// TIA Portal project "1215C_BREAKOUT_BOARD_IO-LINK_TEMPERATURE" (V19)

(* hardware
DEVICE "BREAKOUT_BOARD_PLC"  S7-1200 Station
   slot 0: "Rack_0"  S7-1200 Rack  Rack  V1.0
   slot 1: "BREAKOUT_BOARD_PLC"  CPU 1215C DC/DC/DC  6ES7 215-1AG40-0XB0  V4.6
DEVICE "BREAKOUT_BOARD_HMI"  KTP400 Basic PN
   slot 0: "BREAKOUT_BOARD_HMI"  KTP400 Basic PN  6AV2 123-2DB03-0AX0  16.0.0.0
   slot 1: "HMI_RT_1"  KTP400 Basic PN  6AV2 123-2DB03-0AX0  16.0.0.0
   slot 5: "BREAKOUT_BOARD_HMI.IE_CP_1"  PROFINET Interface  16.0.0.0
      slot 1: "PROFINET Interface"  PROFINET Interface
         slot 1: "Port_1"  Port
DEVICE "IFM_IO-LINK_MASTER"  GSD.Device.PN
   slot 0: "Rack"  Rack  V1.0
   slot 0: "AL1100"  AL1100  AL1100
      slot 0: "AL1100"  AL1100
      slot 1: "X1"  X1
         slot 1: "Port 1"  Port 1
         slot 2: "Port 2"  Port 2
      slot 1: "4 Ports_1"  4 Ports  AL1100
         slot 0: "IO-Link Master"  IO-Link Master
   slot 1: "IFM ITA2105 IO-Link In  2 Byte + PQI"  IO-Link In  2 Byte + PQI
   slot 2: "Disabled_P2"  Disabled
   slot 3: "Disabled_P3"  Disabled
   slot 4: "Disabled_P4"  Disabled
DEVICE "SCALANCE XB008"  SCALANCE X-Station
   slot 0: "SCALANCE X rack"  Rail
   slot 0: "8PORT_SWITCH"  6GK5 008-0BA10-1AB2  V1.0
*)

// ===== PLC "BREAKOUT_BOARD_PLC"  CPU 1215C DC/DC/DC =====

VAR_GLOBAL   // PLC tag table "PLC_Outputs"
   "DQ0.0" AT %Q0.0 : Bool;   // Digital Output
   "DQ0.1" AT %Q0.1 : Bool;   // Digital Output
   "DQ0.2" AT %Q0.2 : Bool;   // Digital Output
   "DQ0.3" AT %Q0.3 : Bool;   // Digital Output
   "DQ0.4" AT %Q0.4 : Bool;   // Digital Output
   "DQ0.5" AT %Q0.5 : Bool;   // Digital Output
   "DQ0.6" AT %Q0.6 : Bool;   // Digital Output
   "DQ0.7" AT %Q0.7 : Bool;   // Digital Output
   "DQ1.0" AT %Q1.0 : Bool;   // Digital Output
   "DQ1.1" AT %Q1.1 : Bool;   // Digital Output
   "AQ0.0" AT %QW64 : Word;   // Analog Output
   "AQ0.1" AT %QW66 : Word;   // Analog Output
END_VAR

VAR_GLOBAL   // PLC tag table "PLC_Inputs"
   "DI0.0" AT %I0.0 : Bool;   // Digital Input
   "DI0.1" AT %I0.1 : Bool;   // Digital Input
   "DI0.2" AT %I0.2 : Bool;   // Digital Input
   "DI0.3" AT %I0.3 : Bool;   // Digital Input
   "DI0.4" AT %I0.4 : Bool;   // Digital Input
   "DI0.5" AT %I0.5 : Bool;   // Digital Input
   "DI0.6" AT %I0.6 : Bool;   // Digital Input
   "DI0.7" AT %I0.7 : Bool;   // Digital Input
   "DI1.0" AT %I1.0 : Bool;   // Digital Input
   "DI1.1" AT %I1.1 : Bool;   // Digital Input
   "DI1.2" AT %I1.2 : Bool;   // Digital Input
   "DI1.3" AT %I1.3 : Bool;   // Digital Input
   "DI1.4" AT %I1.4 : Bool;   // Digital Input
   "DI1.5" AT %I1.5 : Bool;   // Digital Input
   "AI0.0" AT %IW64 : Word;   // Analog Input
   "AI0.1" AT %IW66 : Word;   // Analog Input
END_VAR

VAR_GLOBAL   // PLC tag table "System_Tags"
   "Clock_Byte" AT %MB0 : Byte;
   "Clock_10Hz" AT %M0.0 : Bool;
   "Clock_5Hz" AT %M0.1 : Bool;
   "Clock_2.5Hz" AT %M0.2 : Bool;
   "Clock_2Hz" AT %M0.3 : Bool;
   "Clock_1.25Hz" AT %M0.4 : Bool;
   "Clock_1Hz" AT %M0.5 : Bool;
   "Clock_0.625Hz" AT %M0.6 : Bool;
   "Clock_0.5Hz" AT %M0.7 : Bool;
   "System_Byte" AT %MB1 : Byte;
   "FirstScan" AT %M1.0 : Bool;
   "DiagStatusUpdate" AT %M1.1 : Bool;
   "AlwaysTRUE" AT %M1.2 : Bool;
   "AlwaysFALSE" AT %M1.3 : Bool;
END_VAR

VAR_GLOBAL   // PLC tag table "Trigger_Tags"
   "xAQ_Trig" AT %M2.0 : Bool;
   "xTrig2" AT %M2.1 : Bool;
   "xTrig3" AT %M2.2 : Bool;
   "xTrig4" AT %M2.3 : Bool;
   "xTrig5" AT %M2.4 : Bool;
END_VAR

VAR_GLOBAL   // PLC tag table "IO-Link_Tags"
   "IFM_TA2105_Temp" AT %IW68 : Int;   // IO-Link Master X1
END_VAR

// folder: WS01_TVET_Workstation/00-I/O_Mapping

DATA_BLOCK "DB001-PLC_I/O"   // DB1
TITLE = PLC I/O Global Database
{ S7_Optimized_Access := 'TRUE' }
VERSION : 0.1
// Variables used to mirror the physical PLC I/O states.
   VAR
      Inputs : Struct   // PLC Inputs Structure
         "xDI0.0" : Bool;
         "xDI0.1" : Bool;
         "xDI0.2" : Bool;
         "xDI0.3" : Bool;
         "xDI0.4" : Bool;
         "xDI0.5" : Bool;
         "xDI0.6" : Bool;
         "xDI0.7" : Bool;
         "xDI1.0" : Bool;
         "xDI1.1" : Bool;
         "xDI1.2" : Bool;
         "xDI1.3" : Bool;
         "xDI1.4" : Bool;
         "xDI1.5" : Bool;
         "rAI0.0_Scaled" : Real;   // 0 to 24648 = 0 to 10 V
         "rAI0.1_Scaled" : Real;   // 0 to 24648 = 0 to 10 V
      END_STRUCT;
      Outputs : Struct   // PLC Outputs Structure
         "xDQ0.0" : Bool;
         "xDQ0.1" : Bool;
         "xDQ0.2" : Bool;
         "xDQ0.3" : Bool;
         "xDQ0.4" : Bool;
         "xDQ0.5" : Bool;
         "xDQ0.6" : Bool;
         "xDQ0.7" : Bool;
         "xDQ1.0" : Bool;
         "xDQ1.1" : Bool;
         "iAQ0.0_RAW" : Int := 0;
         "rAQ0.0_Scaled" : Real;   // 0 to 24648 = 0 to 20 mA
         "iAQ0.1_RAW" : Int := 0;
         "rAQ0.1_Scaled" : Real;   // 0 to 24648 = 0 to 20 mA
      END_STRUCT;
   END_VAR
BEGIN
END_DATA_BLOCK

DATA_BLOCK "DB003-IO-Link_I/O"   // DB3
TITLE = IO-Link I/O Global Database
{ S7_Optimized_Access := 'TRUE' }
VERSION : 0.1
// Variables used to mirror the physical IO-Link I/O states.
   VAR
      Inputs : Struct   // IO-Link Inputs Structure
         wTemp_RAW : Word;   // Temperature Sensor Scaled Value
      END_STRUCT;
      Outputs : Struct   // IO-Link Outputs Structure
         wReserved : Word;
      END_STRUCT;
   END_VAR
BEGIN
END_DATA_BLOCK

// folder: WS01_TVET_Workstation/01-Date_Time

DATA_BLOCK "DB002-DateTime"   // DB2
TITLE = PLC Date/Time Global Database
{ S7_Optimized_Access := 'TRUE' }
VERSION : 0.1
// Variables used to store the PLC date/time & custom date/time formatting.
   VAR
      RD_LOC_T_Ret : Int := 0;   // Return value for Read Local Time Block
      LOCAL_DTL : DTL := DTL#1970-01-01-00:00:00;   // RAW DTL
      "Date" : Date := D#1990-01-01;   // RAW Date
      "Time" : Time_Of_Day := TOD#00:00:00;   // RAW Time
      DTLtoString_Ret : String;   // Return value for DTL to String Block
      sCustomDate_YY : String := '';   // Custom year
      sCustomDate_MM : String := '';   // Custom month
      sCustomDate_DD : String := '';   // Custom Day
      sCustomTime_HH : String := '';   // Custom hour
      sCustomTime_MM : String := '';   // Custom minute
      sCustomDate_DDMMYY : String := '';   // Custom date format
      sCustomTime_HHMM : String := '';   // Custom time format
   END_VAR
BEGIN
END_DATA_BLOCK

// folder: WS01_TVET_Workstation/02-IOLink_Control

DATA_BLOCK "DB004-IOLink_Data"   // DB4
TITLE = IO-Link Data Global Database
{ S7_Optimized_Access := 'TRUE' }
VERSION : 0.1
// Variables used to process data from connected devices.
   VAR
      TempSensor_Data : Struct   // Temperature Sensor Data Structure
         rDeg_C : Real;   // Degrees Celsius
         rDeg_F : Real;   // Degrees Fahrenheit
      END_STRUCT;
   END_VAR
BEGIN
END_DATA_BLOCK

// folder: (top level)

ORGANIZATION_BLOCK "Main"   // OB1, LAD, ProgramCycle
TITLE = "Main Program Sweep (Cycle)"
{ S7_Optimized_Access := 'TRUE' }
VERSION : 0.1
   VAR_INPUT
      Initial_Call : Bool;   // Initial call of this OB
      Remanence : Bool;   // =True, if remanent data are available
   END_VAR
BEGIN

REGION Network 1 (SCL): ================= PROGRAM_INFORMATION =================
   (*
   ==================================================================
   ********************* PLC I/O BREAKOUT BOARD *********************
   ==================================================================

   TVET Workstation WS01:
   1215C DC/DC/DC - 6ES7215-1AG40-0XB0 - IP: 192.168.0.175/24

   KTP400 HMI - 6AV2123-2DB03-0AX0 - IP: 192.168.0.176/24

   IFM IO-Link Master - AL1100 - IP: 192.168.0.177/24

   =======================================================================

   The program has 3 main sections:
   - Date/Time Handler,
   - I/O Handlers,
   - IO-Link Devices Handler.

   Date/Time Handler FC:
   - local PLC date/time is read & formatted into a 24HR time & DD/MM/YYYY.

   I/O Handler FCs:
   - maps the physical PLC inputs & outputs to corresponding tags in DB001,
   - handles scaling of the PLC Analog I/O,
   - maps the IO-Link inputs & outputs to corresponding tags in DB003,
   - ensures that physical I/O tags are only used once in the code.

   IO-Link Device Handler FCs:
   - connected IO-Link devices are controlled in this section with the
     temperature sensor conversion logic being handled by an IFM provided
     FC which scales the input value & converts to Fahrenheit.
   - create & call new FC's for any additional IO-Link devices that may
     get added.

   Additional Notes:
   PLC Tags grouped according to their use/function.

   =======================================================================

   Analog Input Technical data:
   - Number of inputs: 2
   - Type: Voltage (single-ended)
   - Full-scale range: 0 to 10 V
   - Full-scale range (data word): 0 to 27648
   - Overshoot range: 10.001 to 11.759 V
   - Overshoot range (data word): 27649 to 32511
   - Overflow range: 11.760 to 11.852 V
   - Overflow range (data word): 32512 to 32767
   - Resolution: 10 bits
   - Maximum withstand voltage: 35 V DC
   - Smoothing: None, Weak, Medium, or Strong
   - Noise rejection: 10, 50, or 60 Hz
   - Impedance: ≥100 KΩ
   - Isolation (field side to logic): None
   - Accuracy (25 °C / -20 to 60 °C): 3.0% / 3.5% of full-scale
   - Cable length (meters): 100 m, shielded twisted pair
   - Rated range: 0     = 0 V
                  34    = 12 mV
                  20736 = 7.5 V
                  27648 = 10 V

   =======================================================================

   Analog Output Technical data:
   - Number of outputs: 2
   - Type: Current
   - Full-scale range: 0 to 20 mA
   - Full-scale range (data word): 0 to 27648
   - Overshoot range: 20.01 to 23.52 mA
   - Overshoot range (data word): 27649 to 32511
   - Overflow range data word: 32512 to 32767
   - Resolution: 10 bits
   - Output drive impedance: ≤500 Ω max
   - Isolation (field side to logic): None
   - Accuracy (25 °C / -20 to 60 °C): 3.0% / 3.5% of full-scale
   - Settling time: 2 ms
   - Cable length (meters): 100 m, shielded twisted pair
   - Rated range: 0     = 0 mA
                  34    = 0.0247 mA
                  20736 = 15 mA
                  27648 = 20 mA

   =======================================================================

   TA2105 IO-Link Temperature Transmitter documentation:
   https://www.ifm.com/us/en/product/TA2105#documents

   Process Data In length = 2bytes

   The IO-Link Inputs screen on the HMI displays a bar graph of the current
   measured temperature for the sensor connected to port X1.

   =======================================================================
   *)
END_REGION

REGION Network 2: ================= LOCAL_DATE/TIME =================
END_REGION

REGION Network 3: Call the Date/Time Handler Function
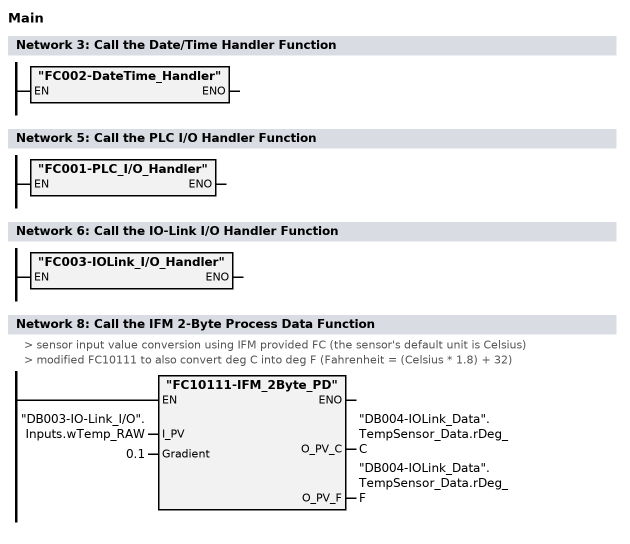
   RUNG wire#powerrail
      "FC002-DateTime_Handler"()
   END_RUNG
   // the same network as SCL:
   "FC002-DateTime_Handler"();
END_REGION

REGION Network 4: ================= I/O_MAPPING =================
END_REGION

REGION Network 5: Call the PLC I/O Handler Function
   RUNG wire#powerrail
      "FC001-PLC_I/O_Handler"()
   END_RUNG
   // the same network as SCL:
   "FC001-PLC_I/O_Handler"();
END_REGION

REGION Network 6: Call the IO-Link I/O Handler Function
   RUNG wire#powerrail
      "FC003-IOLink_I/O_Handler"()
   END_RUNG
   // the same network as SCL:
   "FC003-IOLink_I/O_Handler"();
END_REGION

REGION Network 7: ================= IO-LINK_DEVICES =================
END_REGION

REGION Network 8: Call the IFM 2-Byte Process Data Function
   // > sensor input value conversion using IFM provided FC (the sensor's default unit is Celsius)
   // > modified FC10111 to also convert deg C into deg F (Fahrenheit = (Celsius * 1.8) + 32)
   RUNG wire#powerrail
      "FC10111-IFM_2Byte_PD"(I_PV := "DB003-IO-Link_I/O".Inputs.wTemp_RAW, Gradient := 0.1, O_PV_C => "DB004-IOLink_Data".TempSensor_Data.rDeg_C, O_PV_F => "DB004-IOLink_Data".TempSensor_Data.rDeg_F)
   END_RUNG
   // the same network as SCL:
   "FC10111-IFM_2Byte_PD"(I_PV := "DB003-IO-Link_I/O".Inputs.wTemp_RAW,
                          Gradient := 0.1,
                          O_PV_C => "DB004-IOLink_Data".TempSensor_Data.rDeg_C,
                          O_PV_F => "DB004-IOLink_Data".TempSensor_Data.rDeg_F);
END_REGION
END_ORGANIZATION_BLOCK

// folder: WS01_TVET_Workstation/00-I/O_Mapping

FUNCTION "FC001-PLC_I/O_Handler" : Void   // FC1, LAD
TITLE = PLC Input Output Handler
{ S7_Optimized_Access := 'TRUE' }
VERSION : 0.1
// This function block is for interfacing the physical PLC input/output connections to a Global DB (DB001-PLC_I/O).
   VAR_TEMP
      "rAI0.0_Temp" : Real;
      "rAI0.1_Temp" : Real;
      "rAQ0.0_Temp" : Real;
      "rAQ0.1_Temp" : Real;
   END_VAR
   VAR_TEMP   // added for the SCL form of the ladder/FBD networks
      _w1 : Bool;
   END_VAR
BEGIN

REGION Network 1: ================= DIGITAL_INPUTS =================
END_REGION

REGION Network 2: BANK_0
   // > DI0.0 - DI0.7
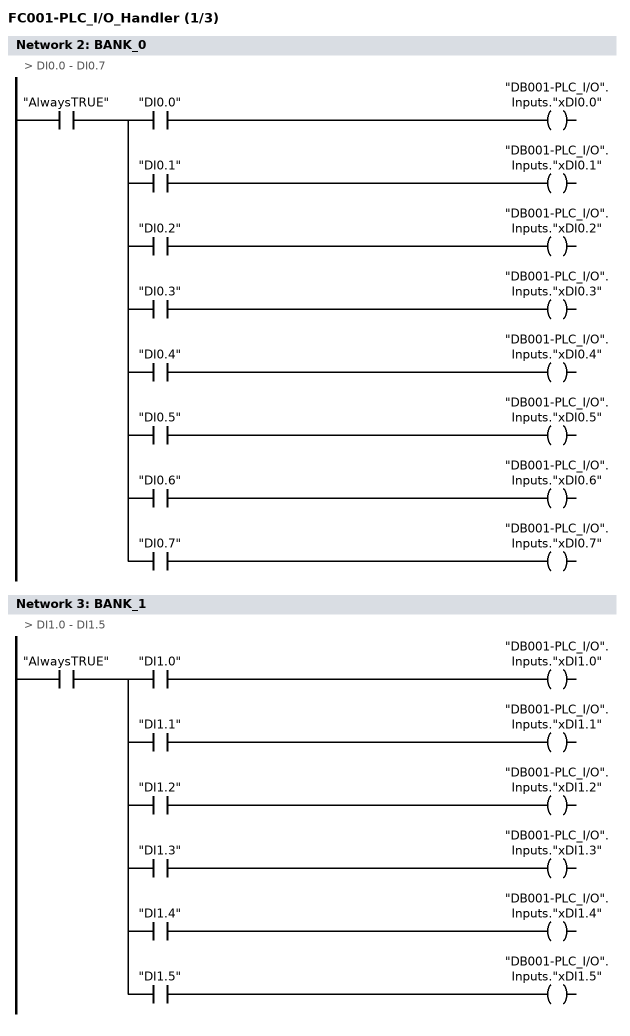
   RUNG wire#powerrail
      Contact( "AlwaysTRUE" )
      wire#w1
      Contact( "DI0.0" )
      Coil( "DB001-PLC_I/O".Inputs."xDI0.0" )
   END_RUNG
   RUNG wire#w1
      Contact( "DI0.1" )
      Coil( "DB001-PLC_I/O".Inputs."xDI0.1" )
   END_RUNG
   RUNG wire#w1
      Contact( "DI0.2" )
      Coil( "DB001-PLC_I/O".Inputs."xDI0.2" )
   END_RUNG
   RUNG wire#w1
      Contact( "DI0.3" )
      Coil( "DB001-PLC_I/O".Inputs."xDI0.3" )
   END_RUNG
   RUNG wire#w1
      Contact( "DI0.4" )
      Coil( "DB001-PLC_I/O".Inputs."xDI0.4" )
   END_RUNG
   RUNG wire#w1
      Contact( "DI0.5" )
      Coil( "DB001-PLC_I/O".Inputs."xDI0.5" )
   END_RUNG
   RUNG wire#w1
      Contact( "DI0.6" )
      Coil( "DB001-PLC_I/O".Inputs."xDI0.6" )
   END_RUNG
   RUNG wire#w1
      Contact( "DI0.7" )
      Coil( "DB001-PLC_I/O".Inputs."xDI0.7" )
   END_RUNG
   // the same network as SCL:
   "DB001-PLC_I/O".Inputs."xDI0.0" := "AlwaysTRUE" AND "DI0.0";
   "DB001-PLC_I/O".Inputs."xDI0.1" := "AlwaysTRUE" AND "DI0.1";
   "DB001-PLC_I/O".Inputs."xDI0.2" := "AlwaysTRUE" AND "DI0.2";
   "DB001-PLC_I/O".Inputs."xDI0.3" := "AlwaysTRUE" AND "DI0.3";
   "DB001-PLC_I/O".Inputs."xDI0.4" := "AlwaysTRUE" AND "DI0.4";
   "DB001-PLC_I/O".Inputs."xDI0.5" := "AlwaysTRUE" AND "DI0.5";
   "DB001-PLC_I/O".Inputs."xDI0.6" := "AlwaysTRUE" AND "DI0.6";
   "DB001-PLC_I/O".Inputs."xDI0.7" := "AlwaysTRUE" AND "DI0.7";
END_REGION

REGION Network 3: BANK_1
   // > DI1.0 - DI1.5
   RUNG wire#powerrail
      Contact( "AlwaysTRUE" )
      wire#w1
      Contact( "DI1.0" )
      Coil( "DB001-PLC_I/O".Inputs."xDI1.0" )
   END_RUNG
   RUNG wire#w1
      Contact( "DI1.1" )
      Coil( "DB001-PLC_I/O".Inputs."xDI1.1" )
   END_RUNG
   RUNG wire#w1
      Contact( "DI1.2" )
      Coil( "DB001-PLC_I/O".Inputs."xDI1.2" )
   END_RUNG
   RUNG wire#w1
      Contact( "DI1.3" )
      Coil( "DB001-PLC_I/O".Inputs."xDI1.3" )
   END_RUNG
   RUNG wire#w1
      Contact( "DI1.4" )
      Coil( "DB001-PLC_I/O".Inputs."xDI1.4" )
   END_RUNG
   RUNG wire#w1
      Contact( "DI1.5" )
      Coil( "DB001-PLC_I/O".Inputs."xDI1.5" )
   END_RUNG
   // the same network as SCL:
   "DB001-PLC_I/O".Inputs."xDI1.0" := "AlwaysTRUE" AND "DI1.0";
   "DB001-PLC_I/O".Inputs."xDI1.1" := "AlwaysTRUE" AND "DI1.1";
   "DB001-PLC_I/O".Inputs."xDI1.2" := "AlwaysTRUE" AND "DI1.2";
   "DB001-PLC_I/O".Inputs."xDI1.3" := "AlwaysTRUE" AND "DI1.3";
   "DB001-PLC_I/O".Inputs."xDI1.4" := "AlwaysTRUE" AND "DI1.4";
   "DB001-PLC_I/O".Inputs."xDI1.5" := "AlwaysTRUE" AND "DI1.5";
END_REGION

REGION Network 4: ================= DIGITAL_OUTPUTS =================
END_REGION

REGION Network 5: BANK_0
   // > DQ0.0 - DQ0.7
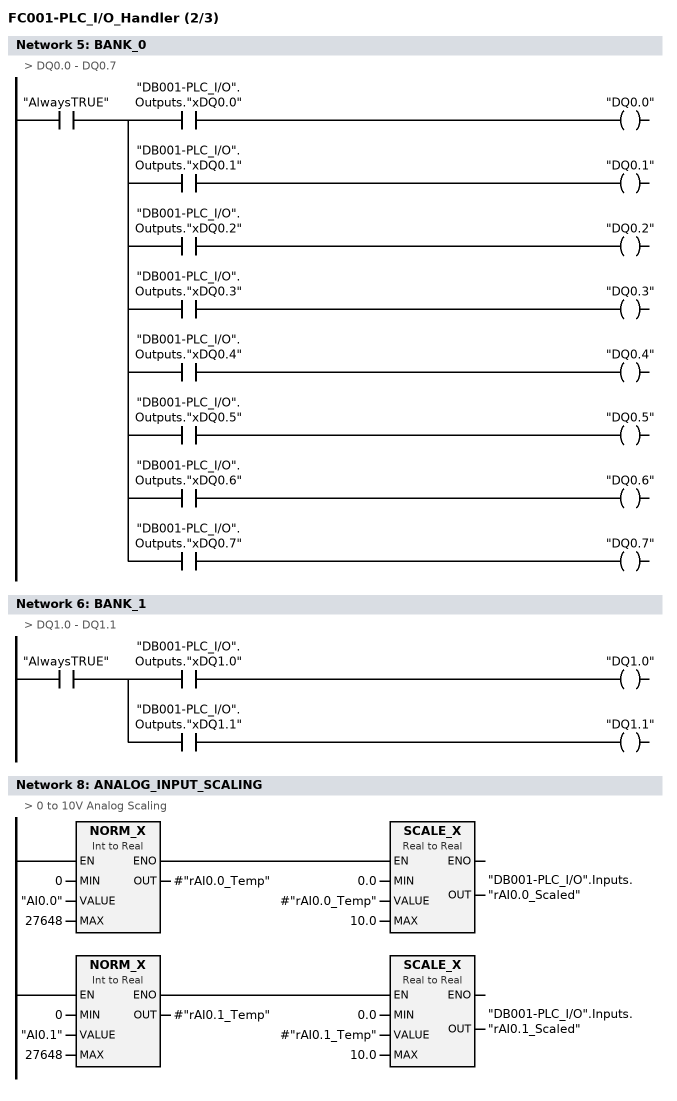
   RUNG wire#powerrail
      Contact( "AlwaysTRUE" )
      wire#w1
      Contact( "DB001-PLC_I/O".Outputs."xDQ0.0" )
      Coil( "DQ0.0" )
   END_RUNG
   RUNG wire#w1
      Contact( "DB001-PLC_I/O".Outputs."xDQ0.1" )
      Coil( "DQ0.1" )
   END_RUNG
   RUNG wire#w1
      Contact( "DB001-PLC_I/O".Outputs."xDQ0.2" )
      Coil( "DQ0.2" )
   END_RUNG
   RUNG wire#w1
      Contact( "DB001-PLC_I/O".Outputs."xDQ0.3" )
      Coil( "DQ0.3" )
   END_RUNG
   RUNG wire#w1
      Contact( "DB001-PLC_I/O".Outputs."xDQ0.4" )
      Coil( "DQ0.4" )
   END_RUNG
   RUNG wire#w1
      Contact( "DB001-PLC_I/O".Outputs."xDQ0.5" )
      Coil( "DQ0.5" )
   END_RUNG
   RUNG wire#w1
      Contact( "DB001-PLC_I/O".Outputs."xDQ0.6" )
      Coil( "DQ0.6" )
   END_RUNG
   RUNG wire#w1
      Contact( "DB001-PLC_I/O".Outputs."xDQ0.7" )
      Coil( "DQ0.7" )
   END_RUNG
   // the same network as SCL:
   "DQ0.0" := "AlwaysTRUE" AND "DB001-PLC_I/O".Outputs."xDQ0.0";
   "DQ0.1" := "AlwaysTRUE" AND "DB001-PLC_I/O".Outputs."xDQ0.1";
   "DQ0.2" := "AlwaysTRUE" AND "DB001-PLC_I/O".Outputs."xDQ0.2";
   "DQ0.3" := "AlwaysTRUE" AND "DB001-PLC_I/O".Outputs."xDQ0.3";
   "DQ0.4" := "AlwaysTRUE" AND "DB001-PLC_I/O".Outputs."xDQ0.4";
   "DQ0.5" := "AlwaysTRUE" AND "DB001-PLC_I/O".Outputs."xDQ0.5";
   "DQ0.6" := "AlwaysTRUE" AND "DB001-PLC_I/O".Outputs."xDQ0.6";
   "DQ0.7" := "AlwaysTRUE" AND "DB001-PLC_I/O".Outputs."xDQ0.7";
END_REGION

REGION Network 6: BANK_1
   // > DQ1.0 - DQ1.1
   RUNG wire#powerrail
      Contact( "AlwaysTRUE" )
      wire#w1
      Contact( "DB001-PLC_I/O".Outputs."xDQ1.0" )
      Coil( "DQ1.0" )
   END_RUNG
   RUNG wire#w1
      Contact( "DB001-PLC_I/O".Outputs."xDQ1.1" )
      Coil( "DQ1.1" )
   END_RUNG
   // the same network as SCL:
   "DQ1.0" := "AlwaysTRUE" AND "DB001-PLC_I/O".Outputs."xDQ1.0";
   "DQ1.1" := "AlwaysTRUE" AND "DB001-PLC_I/O".Outputs."xDQ1.1";
END_REGION

REGION Network 7: ================= ANALOG_PROCESSING =================
END_REGION

REGION Network 8: ANALOG_INPUT_SCALING
   // > 0 to 10V Analog Scaling
   RUNG wire#powerrail
      { S7_Templates := "[SrcType := Int, DestType := Real]" } Normalize(min := 0, value := "AI0.0", max := 27648, out => #"rAI0.0_Temp")
      { S7_Templates := "[SrcType := Real, DestType := Real]" } Scale(min := 0.0, value := #"rAI0.0_Temp", max := 10.0, out => "DB001-PLC_I/O".Inputs."rAI0.0_Scaled")
   END_RUNG
   RUNG wire#powerrail
      { S7_Templates := "[SrcType := Int, DestType := Real]" } Normalize(min := 0, value := "AI0.1", max := 27648, out => #"rAI0.1_Temp")
      { S7_Templates := "[SrcType := Real, DestType := Real]" } Scale(min := 0.0, value := #"rAI0.1_Temp", max := 10.0, out => "DB001-PLC_I/O".Inputs."rAI0.1_Scaled")
   END_RUNG
   // the same network as SCL:
   #"rAI0.0_Temp" := NORM_X(MIN := 0, VALUE := "AI0.0", MAX := 27648);
   "DB001-PLC_I/O".Inputs."rAI0.0_Scaled" := SCALE_X(MIN := 0.0, VALUE := #"rAI0.0_Temp", MAX := 10.0);
   #"rAI0.1_Temp" := NORM_X(MIN := 0, VALUE := "AI0.1", MAX := 27648);
   "DB001-PLC_I/O".Inputs."rAI0.1_Scaled" := SCALE_X(MIN := 0.0, VALUE := #"rAI0.1_Temp", MAX := 10.0);
END_REGION

REGION Network 9: ANALOG_OUTPUT_SCALING
   // > 0 to 20mA Analog Scaling
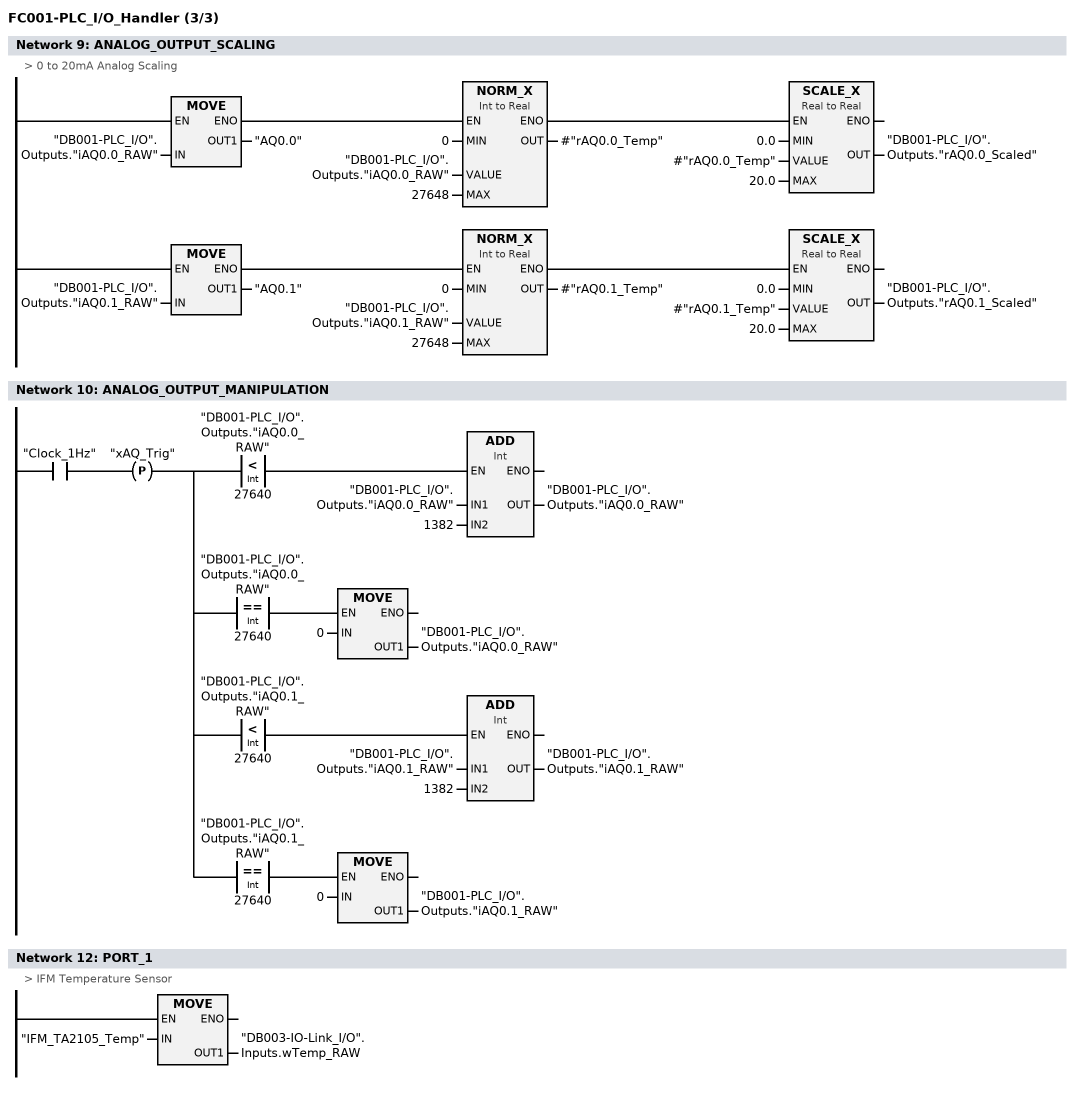
   RUNG wire#powerrail
      Move(in := "DB001-PLC_I/O".Outputs."iAQ0.0_RAW", out1 => "AQ0.0")
      { S7_Templates := "[SrcType := Int, DestType := Real]" } Normalize(min := 0, value := "DB001-PLC_I/O".Outputs."iAQ0.0_RAW", max := 27648, out => #"rAQ0.0_Temp")
      { S7_Templates := "[SrcType := Real, DestType := Real]" } Scale(min := 0.0, value := #"rAQ0.0_Temp", max := 20.0, out => "DB001-PLC_I/O".Outputs."rAQ0.0_Scaled")
   END_RUNG
   RUNG wire#powerrail
      Move(in := "DB001-PLC_I/O".Outputs."iAQ0.1_RAW", out1 => "AQ0.1")
      { S7_Templates := "[SrcType := Int, DestType := Real]" } Normalize(min := 0, value := "DB001-PLC_I/O".Outputs."iAQ0.1_RAW", max := 27648, out => #"rAQ0.1_Temp")
      { S7_Templates := "[SrcType := Real, DestType := Real]" } Scale(min := 0.0, value := #"rAQ0.1_Temp", max := 20.0, out => "DB001-PLC_I/O".Outputs."rAQ0.1_Scaled")
   END_RUNG
   // the same network as SCL:
   "AQ0.0" := "DB001-PLC_I/O".Outputs."iAQ0.0_RAW";
   #"rAQ0.0_Temp" := NORM_X(MIN := 0, VALUE := "DB001-PLC_I/O".Outputs."iAQ0.0_RAW", MAX := 27648);
   "DB001-PLC_I/O".Outputs."rAQ0.0_Scaled" := SCALE_X(MIN := 0.0, VALUE := #"rAQ0.0_Temp", MAX := 20.0);
   "AQ0.1" := "DB001-PLC_I/O".Outputs."iAQ0.1_RAW";
   #"rAQ0.1_Temp" := NORM_X(MIN := 0, VALUE := "DB001-PLC_I/O".Outputs."iAQ0.1_RAW", MAX := 27648);
   "DB001-PLC_I/O".Outputs."rAQ0.1_Scaled" := SCALE_X(MIN := 0.0, VALUE := #"rAQ0.1_Temp", MAX := 20.0);
END_REGION

REGION Network 10: ANALOG_OUTPUT_MANIPULATION
   RUNG wire#powerrail
      Contact( "Clock_1Hz" )
      P_Trig( "xAQ_Trig" )
      wire#w1
      { S7_Templates := "SrcType := Int" } LT_Contact(in1 := "DB001-PLC_I/O".Outputs."iAQ0.0_RAW", in2 := 27640)
      { S7_Templates := "SrcType := Int" } Add(in1 := "DB001-PLC_I/O".Outputs."iAQ0.0_RAW", in2 := 1382, out => "DB001-PLC_I/O".Outputs."iAQ0.0_RAW")
   END_RUNG
   RUNG wire#w1
      { S7_Templates := "SrcType := Int" } EQ_Contact(in1 := "DB001-PLC_I/O".Outputs."iAQ0.0_RAW", in2 := 27640)
      Move(in := 0, out1 => "DB001-PLC_I/O".Outputs."iAQ0.0_RAW")
   END_RUNG
   RUNG wire#w1
      { S7_Templates := "SrcType := Int" } LT_Contact(in1 := "DB001-PLC_I/O".Outputs."iAQ0.1_RAW", in2 := 27640)
      { S7_Templates := "SrcType := Int" } Add(in1 := "DB001-PLC_I/O".Outputs."iAQ0.1_RAW", in2 := 1382, out => "DB001-PLC_I/O".Outputs."iAQ0.1_RAW")
   END_RUNG
   RUNG wire#w1
      { S7_Templates := "SrcType := Int" } EQ_Contact(in1 := "DB001-PLC_I/O".Outputs."iAQ0.1_RAW", in2 := 27640)
      Move(in := 0, out1 => "DB001-PLC_I/O".Outputs."iAQ0.1_RAW")
   END_RUNG
   // the same network as SCL:
   #_w1 := "Clock_1Hz" AND NOT "xAQ_Trig";   // rising edge
   "xAQ_Trig" := "Clock_1Hz";
   IF #_w1 AND ("DB001-PLC_I/O".Outputs."iAQ0.0_RAW" < 27640) THEN
       "DB001-PLC_I/O".Outputs."iAQ0.0_RAW" := "DB001-PLC_I/O".Outputs."iAQ0.0_RAW" + 1382;
   END_IF;
   IF #_w1 AND ("DB001-PLC_I/O".Outputs."iAQ0.0_RAW" = 27640) THEN
       "DB001-PLC_I/O".Outputs."iAQ0.0_RAW" := 0;
   END_IF;
   IF #_w1 AND ("DB001-PLC_I/O".Outputs."iAQ0.1_RAW" < 27640) THEN
       "DB001-PLC_I/O".Outputs."iAQ0.1_RAW" := "DB001-PLC_I/O".Outputs."iAQ0.1_RAW" + 1382;
   END_IF;
   IF #_w1 AND ("DB001-PLC_I/O".Outputs."iAQ0.1_RAW" = 27640) THEN
       "DB001-PLC_I/O".Outputs."iAQ0.1_RAW" := 0;
   END_IF;
END_REGION

REGION Network 11: ================= IO-LINK_INPUTS =================
END_REGION

REGION Network 12: PORT_1
   // > IFM Temperature Sensor
   RUNG wire#powerrail
      Move(in := "IFM_TA2105_Temp", out1 => "DB003-IO-Link_I/O".Inputs.wTemp_RAW)
   END_RUNG
   // the same network as SCL:
   "DB003-IO-Link_I/O".Inputs.wTemp_RAW := "IFM_TA2105_Temp";
END_REGION

REGION Network 13: ================= IO-LINK_OUTPUTS =================
END_REGION

REGION Network 14: PORT_2
END_REGION
END_FUNCTION

FUNCTION "FC003-IOLink_I/O_Handler" : Void   // FC3, LAD
TITLE = IOLink Input/Output Handler
{ S7_Optimized_Access := 'TRUE' }
VERSION : 0.1
// This function block is for interfacing the physical IO-Link input/output data to a Global DB (DB003-IOLink_I/O).
BEGIN

REGION Network 1: ================= PORT_X1 =================
END_REGION

REGION Network 2: IFM Temperature Sensor
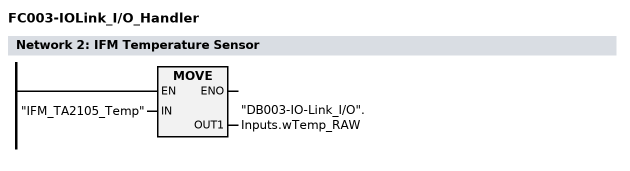
   RUNG wire#powerrail
      Move(in := "IFM_TA2105_Temp", out1 => "DB003-IO-Link_I/O".Inputs.wTemp_RAW)
   END_RUNG
   // the same network as SCL:
   "DB003-IO-Link_I/O".Inputs.wTemp_RAW := "IFM_TA2105_Temp";
END_REGION

REGION Network 3: ================= PORT_X2 =================
END_REGION

REGION Network 4: Reserved
END_REGION
END_FUNCTION

// folder: WS01_TVET_Workstation/01-Date_Time

FUNCTION "FC002-DateTime_Handler" : Void   // FC2, LAD
TITLE = Date Time Handler
{ S7_Optimized_Access := 'TRUE' }
VERSION : 0.1
// This function block is for formatting the PLC time into a format suitable for display on the HMI.
   VAR_TEMP   // added for the SCL form of the ladder/FBD networks
      _w1 : Bool;
   END_VAR
BEGIN

REGION Network 1: Read Local Date/Time
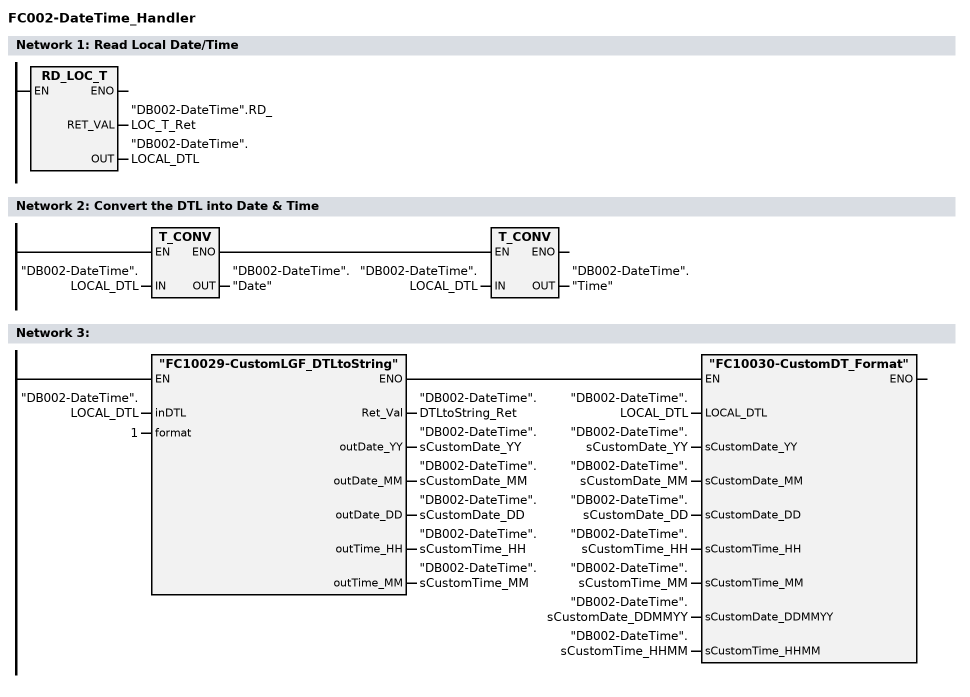
   "DB002-DateTime".RD_LOC_T_Ret := RD_LOC_T(OUT => "DB002-DateTime".LOCAL_DTL);
END_REGION

REGION Network 2: Convert the DTL into Date & Time
   // ENO of a box is taken as its EN; it also drops when the box reports an error
   "DB002-DateTime"."Date" := T_CONV(IN := "DB002-DateTime".LOCAL_DTL);
   "DB002-DateTime"."Time" := T_CONV(IN := "DB002-DateTime".LOCAL_DTL);
END_REGION

REGION Network 3
   RUNG wire#powerrail
      "FC10029-CustomLGF_DTLtoString"(inDTL := "DB002-DateTime".LOCAL_DTL, format := 1, Ret_Val => "DB002-DateTime".DTLtoString_Ret, outDate_YY => "DB002-DateTime".sCustomDate_YY, outDate_MM => "DB002-DateTime".sCustomDate_MM, outDate_DD => "DB002-DateTime".sCustomDate_DD, outTime_HH => "DB002-DateTime".sCustomTime_HH, outTime_MM => "DB002-DateTime".sCustomTime_MM)
      "FC10030-CustomDT_Format"(LOCAL_DTL := "DB002-DateTime".LOCAL_DTL, sCustomDate_YY := "DB002-DateTime".sCustomDate_YY, sCustomDate_MM := "DB002-DateTime".sCustomDate_MM, sCustomDate_DD := "DB002-DateTime".sCustomDate_DD, sCustomTime_HH := "DB002-DateTime".sCustomTime_HH, sCustomTime_MM := "DB002-DateTime".sCustomTime_MM, sCustomDate_DDMMYY := "DB002-DateTime".sCustomDate_DDMMYY, sCustomTime_HHMM := "DB002-DateTime".sCustomTime_HHMM)
   END_RUNG
   // the same network as SCL:
   "DB002-DateTime".DTLtoString_Ret := "FC10029-CustomLGF_DTLtoString"(inDTL := "DB002-DateTime".LOCAL_DTL,
                           format := 1,
                           outDate_YY => "DB002-DateTime".sCustomDate_YY,
                           outDate_MM => "DB002-DateTime".sCustomDate_MM,
                           outDate_DD => "DB002-DateTime".sCustomDate_DD,
                           outTime_HH => "DB002-DateTime".sCustomTime_HH,
                           outTime_MM => "DB002-DateTime".sCustomTime_MM,
                           ENO => #_w1);
   IF #_w1 THEN
       "FC10030-CustomDT_Format"(LOCAL_DTL := "DB002-DateTime".LOCAL_DTL,
                               sCustomDate_YY := "DB002-DateTime".sCustomDate_YY,
                               sCustomDate_MM := "DB002-DateTime".sCustomDate_MM,
                               sCustomDate_DD := "DB002-DateTime".sCustomDate_DD,
                               sCustomTime_HH := "DB002-DateTime".sCustomTime_HH,
                               sCustomTime_MM := "DB002-DateTime".sCustomTime_MM,
                               sCustomDate_DDMMYY := "DB002-DateTime".sCustomDate_DDMMYY,
                               sCustomTime_HHMM := "DB002-DateTime".sCustomTime_HHMM);
   END_IF;
END_REGION
END_FUNCTION

FUNCTION "FC10029-CustomLGF_DTLtoString" : String   // FC10029, SCL
TITLE = Custom LGF Local Date TIme to String Converter
{ S7_Optimized_Access := 'TRUE' }
VERSION : 0.1
// This function block is a modified version of the DTLtoString FC provided by Siemens in the LGF Library.
   VAR_INPUT
      inDTL : DTL;   // Date as DTL tag
      format : Bool;   // 1 = traditional, 0 = international
   END_VAR
   VAR_OUTPUT
      outDate_YY : String;   // Custom Date Output (YY)
      outDate_MM : String;   // Custom Date Output (MM)
      outDate_DD : String;   // Custom Date Output (DD)
      outTime_HH : String;   // Custom Time Output (HH)
      outTime_MM : String;   // Custom Time Output (MM)
   END_VAR
   VAR_TEMP
      tempString : String;   // -
      tempSepTime : Char;   // -
      tempPosYear : USInt;   // -
      tempPosMonth : USInt;   // -
      tempPosDay : USInt;   // -
      tempPosHour : USInt;   // -
      tempPosMinute : USInt;   // -
      tempPosSepYearMonth : USInt;   // -
      tempPosSepMonthDay : USInt;   // -
      tempPosSepHourMinute : USInt;   // -
   END_VAR
   // Ret_Val : Date as String tag
BEGIN
   //=============================================================================
   // Siemens AG
   // (c)Copyright 2017
   //-----------------------------------------------------------------------------
   // Library:       LGF (Library General Functions)
   // Tested with:   CPU1212C DC/DC/DC FW:V4.2
   // Engineering:   TIA Portal V14 Update 1
   // Restrictions:  -
   // Requirements:  PLC (S7-1200 / S7-1500)
   // Functionality: This function converts DTL into a string.  (EDITED)
   //-----------------------------------------------------------------------------
   // Change log table:
   // Version  Date        In charge / Changes applied
   // 01.00.00 15.06.2016  Siemens Industry Online Support
   //                      First released version
   // 01.00.01 02.01.2017  Siemens Industry Online Support
   //                      Upgrade: TIA Portal V14 Update 1
   // 01.00.02 17.08.2018  Siemens Industry Online Support
   //                      Upgrade: TIA V15 Update 2
   //=============================================================================


   // Initialization
   #tempString := '';
   #tempSepTime := ':';


   // Set format parameters for output string
   IF NOT #format
   THEN                                          // International ISO 8601
       #tempPosYear := 1;                          // DTL  | Y| Y| Y| Y| -| M| M| -| D| D|  | H| H| :| M| M|
       #tempPosMonth := 6;                         // -----|--|--|--|--|--|--|--|--|--|--|--|--|--|--|--|--|
       #tempPosDay := 9;                           // Pos  | 1| 2| 3| 4| 5| 6| 7| 8| 9|10|11|12|13|14|15|16|
       #tempPosHour := 12;
       #tempPosMinute := 15;
       #tempPosSepYearMonth := 5;
       #tempPosSepMonthDay := 8;
       #tempPosSepHourMinute := 14;
   ELSE                                          // Traditional (EU)
       #tempPosYear := 7;                          // DTL  | D| D| -| M| M| -| Y| Y| Y| Y|  | H| H| :| M| M|
       #tempPosMonth := 4;                         // -----|--|--|--|--|--|--|--|--|--|--|--|--|--|--|--|--|
       #tempPosDay := 1;                           // Pos  | 1| 2| 3| 4| 5| 6| 7| 8| 9|10|11|12|13|14|15|16|
       #tempPosHour := 12;
       #tempPosMinute := 15;
       #tempPosSepYearMonth := 6;
       #tempPosSepMonthDay := 3;
       #tempPosSepHourMinute := 14;
   END_IF;


   // Convert "Value" into "String" and place at the right position

   // Convert for YEAR
   VAL_STRG(FORMAT := W#16#0000,
            IN := #inDTL.YEAR,
            P := #tempPosYear,
            PREC := 0,
            SIZE := 4,
            OUT => #tempString);     // DTL YEAR --> String --> #tempPosYear

   VAL_STRG(FORMAT := W#16#0000,
            IN := #inDTL.YEAR MOD 100,
            P := 1,
            PREC := 0,
            SIZE := 2,
            OUT => #outDate_YY);        // DTL YEAR --> String --> #CustOutYear (Last 2 digits)

   // Convert for MONTH
   VAL_STRG(FORMAT := W#16#0000,
            IN := #inDTL.MONTH,
            P := #tempPosMonth,
            PREC := 0,
            SIZE := 2,
            OUT => #tempString);     // DTL MONTH --> String --> #tempPosMonth

   VAL_STRG(FORMAT := W#16#0000,
            IN := #inDTL.MONTH,
            P := 1,
            PREC := 0,
            SIZE := 2,
            OUT => #outDate_MM);        // DTL MONTH --> String --> #CustOutDate MM

   // Convert for DAY
   VAL_STRG(FORMAT := W#16#0000,
            IN := #inDTL.DAY,
            P := #tempPosDay,
            PREC := 0,
            SIZE := 2,
            OUT => #tempString);     // DTL DAY --> String --> #tempPosDay

   VAL_STRG(FORMAT := W#16#0000,
            IN := #inDTL.DAY,
            P := 1,
            PREC := 0,
            SIZE := 2,
            OUT => #outDate_DD);        // DTL DAY --> String --> #CustOutDate DDMM

   // Convert for HOUR
   VAL_STRG(FORMAT := W#16#0000,
            IN := #inDTL.HOUR,
            P := #tempPosHour,
            PREC := 0,
            SIZE := 2,
            OUT => #tempString);     // DTL HOUR --> String --> #tempPosHour

   VAL_STRG(FORMAT := W#16#0000,
            IN := #inDTL.HOUR,
            P := 1,
            PREC := 0,
            SIZE := 2,
            OUT => #outTime_HH);     // DTL HOUR --> String --> #CustOutTime HH

   // Convert for MINUTE
   VAL_STRG(FORMAT := W#16#0000,
            IN := #inDTL.MINUTE,
            P := #tempPosMinute,
            PREC := 0,
            SIZE := 2,
            OUT => #tempString);     // DTL MINUTE --> String --> #tempPosMinute

   VAL_STRG(FORMAT := W#16#0000,
            IN := #inDTL.MINUTE,
            P := 1,
            PREC := 0,
            SIZE := 2,
            OUT => #outTime_MM);        // DTL MINUTE --> String --> #CustOutTime


   // Block output
   #"FC10029-CustomLGF_DTLtoString" := #tempString;


   // Additional outputs
   #outDate_YY := #outDate_YY;
   #outDate_MM := #outDate_MM;
   #outDate_DD := #outDate_DD;
   #outTime_HH := #outTime_HH;
   #outTime_MM := #outTime_MM;
END_FUNCTION

FUNCTION "FC10030-CustomDT_Format" : Void   // FC10030, LAD
TITLE = Custom Date/Time Formats
{ S7_Optimized_Access := 'TRUE' }
VERSION : 0.1
// This function block is for formatting the local date/time display on the HMI.
   VAR_INPUT
      LOCAL_DTL : DTL;   // RAW DTL
   END_VAR
   VAR_IN_OUT
      sCustomDate_YY : String;   // Custom Year Output (YY)
      sCustomDate_MM : String;   // Custom Date Output (MM)
      sCustomDate_DD : String;   // Custom Date Output (DD)
      sCustomTime_HH : String;   // Custom Time Output (HH)
      sCustomTime_MM : String;   // Custom Time Output (MM)
      sCustomDate_DDMMYY : String;   // Custom Date (DD/MM/YY)
      sCustomTime_HHMM : String;   // Custom Date (HH:MM)
   END_VAR
   VAR_TEMP
      sTemp_String : String;   // -
   END_VAR
BEGIN

REGION Network 1: =================ADD_LEADING_ZEROS=================
END_REGION

REGION Network 2: Add leading zero to MM if less than 10
   // > If DTL.MONTH is less than 10 - replace 1st character in DD with a 0
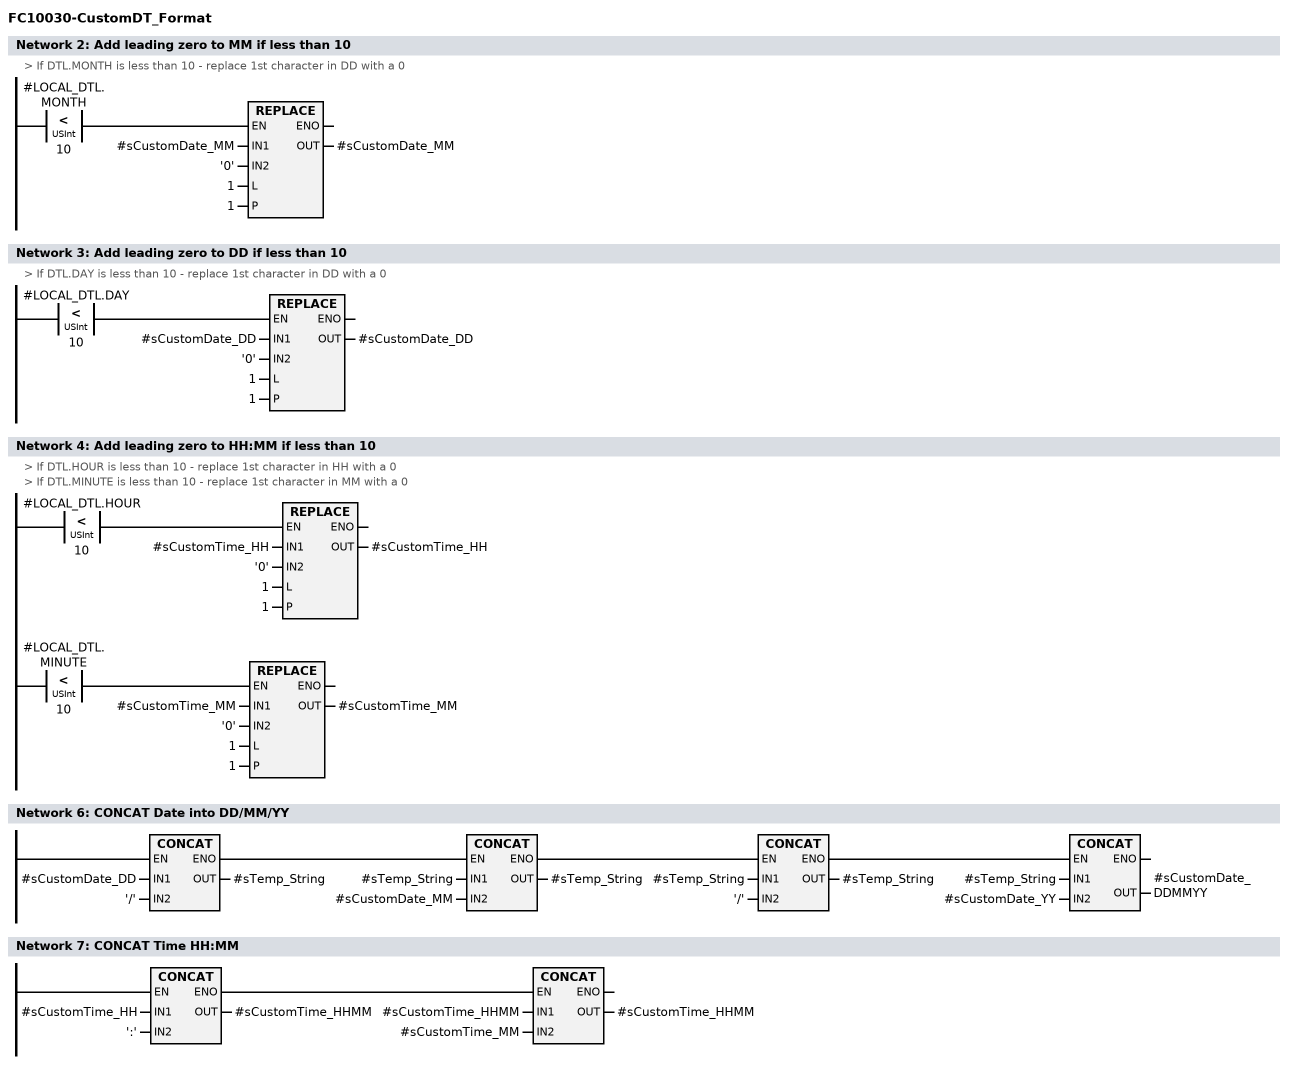
   IF #LOCAL_DTL.MONTH < 10 THEN
       #sCustomDate_MM := REPLACE(IN1 := #sCustomDate_MM, IN2 := '0', L := 1, P := 1);
   END_IF;
END_REGION

REGION Network 3: Add leading zero to DD if less than 10
   // > If DTL.DAY is less than 10 - replace 1st character in DD with a 0
   IF #LOCAL_DTL.DAY < 10 THEN
       #sCustomDate_DD := REPLACE(IN1 := #sCustomDate_DD, IN2 := '0', L := 1, P := 1);
   END_IF;
END_REGION
